// TIA Portal project "Tes simulation extract_V15.1" (V15.1) (continued)
VERSION : 0.1
   VAR_TEMP   // added for the SCL form of the ladder/FBD networks
      _w1 : Bool;
      _w2 : Bool;
   END_VAR
BEGIN

REGION Network 1: BUKA VALVE VP 1 DAN VP 5
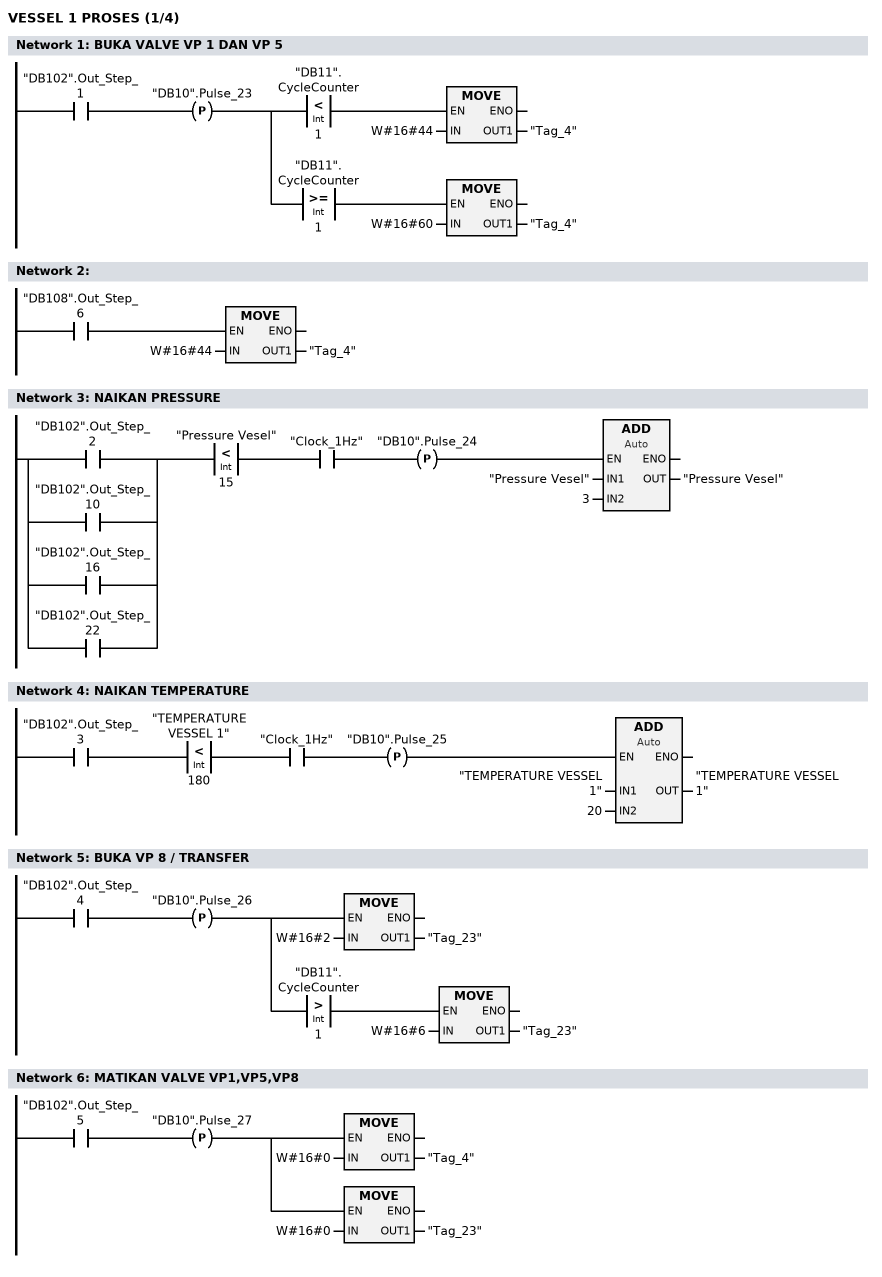
   RUNG wire#powerrail
      Contact( "DB102".Out_Step_1 )
      P_Trig( "DB10".Pulse_23 )
      wire#w1
      { S7_Templates := "SrcType := Int" } LT_Contact(in1 := "DB11".CycleCounter, in2 := 1)
      Move(in := W#16#44, out1 => "Tag_4")
   END_RUNG
   RUNG wire#w1
      { S7_Templates := "SrcType := Int" } GE_Contact(in1 := "DB11".CycleCounter, in2 := 1)
      Move(in := W#16#60, out1 => "Tag_4")
   END_RUNG
   // the same network as SCL:
   #_w1 := "DB102".Out_Step_1 AND NOT "DB10".Pulse_23;   // rising edge
   "DB10".Pulse_23 := "DB102".Out_Step_1;
   IF #_w1 AND ("DB11".CycleCounter < 1) THEN "Tag_4" := W#16#44; END_IF;
   IF #_w1 AND ("DB11".CycleCounter >= 1) THEN "Tag_4" := W#16#60; END_IF;
END_REGION

REGION Network 2
   RUNG wire#powerrail
      Contact( "DB108".Out_Step_6 )
      Move(in := W#16#44, out1 => "Tag_4")
   END_RUNG
   // the same network as SCL:
   IF "DB108".Out_Step_6 THEN "Tag_4" := W#16#44; END_IF;
END_REGION

REGION Network 3: NAIKAN PRESSURE
   RUNG wire#powerrail
      Contact( "DB102".Out_Step_2 )
      wire#w1
      { S7_Templates := "SrcType := Int" } LT_Contact(in1 := "Pressure Vesel", in2 := 15)
      Contact( "Clock_1Hz" )
      P_Trig( "DB10".Pulse_24 )
      Add(in1 := "Pressure Vesel", in2 := 3, out => "Pressure Vesel")
   END_RUNG
   RUNG wire#powerrail
      Contact( "DB102".Out_Step_10 )
   END_RUNG wire#w1
   RUNG wire#powerrail
      Contact( "DB102".Out_Step_16 )
   END_RUNG wire#w1
   RUNG wire#powerrail
      Contact( "DB102".Out_Step_22 )
   END_RUNG wire#w1
   // the same network as SCL:
   #_w1 := ("DB102".Out_Step_2 OR "DB102".Out_Step_10 OR "DB102".Out_Step_16 OR "DB102".Out_Step_22) AND ("Pressure Vesel" < 15) AND "Clock_1Hz";
   #_w2 := #_w1 AND NOT "DB10".Pulse_24;   // rising edge
   "DB10".Pulse_24 := #_w1;
   IF #_w2 THEN "Pressure Vesel" := "Pressure Vesel" + 3; END_IF;
END_REGION

REGION Network 4: NAIKAN TEMPERATURE
   RUNG wire#powerrail
      Contact( "DB102".Out_Step_3 )
      { S7_Templates := "SrcType := Int" } LT_Contact(in1 := "TEMPERATURE VESSEL 1", in2 := 180)
      Contact( "Clock_1Hz" )
      P_Trig( "DB10".Pulse_25 )
      Add(in1 := "TEMPERATURE VESSEL 1", in2 := 20, out => "TEMPERATURE VESSEL 1")
   END_RUNG
   // the same network as SCL:
   #_w1 := "DB102".Out_Step_3 AND ("TEMPERATURE VESSEL 1" < 180) AND "Clock_1Hz";
   #_w2 := #_w1 AND NOT "DB10".Pulse_25;   // rising edge
   "DB10".Pulse_25 := #_w1;
   IF #_w2 THEN "TEMPERATURE VESSEL 1" := "TEMPERATURE VESSEL 1" + 20; END_IF;
END_REGION

REGION Network 5: BUKA VP 8 / TRANSFER
   RUNG wire#powerrail
      Contact( "DB102".Out_Step_4 )
      P_Trig( "DB10".Pulse_26 )
      wire#w1
      Move(in := W#16#2, out1 => "Tag_23")
   END_RUNG
   RUNG wire#w1
      { S7_Templates := "SrcType := Int" } GT_Contact(in1 := "DB11".CycleCounter, in2 := 1)
      Move(in := W#16#6, out1 => "Tag_23")
   END_RUNG
   // the same network as SCL:
   #_w1 := "DB102".Out_Step_4 AND NOT "DB10".Pulse_26;   // rising edge
   "DB10".Pulse_26 := "DB102".Out_Step_4;
   IF #_w1 THEN "Tag_23" := W#16#2; END_IF;
   IF #_w1 AND ("DB11".CycleCounter > 1) THEN "Tag_23" := W#16#6; END_IF;
END_REGION

REGION Network 6: MATIKAN VALVE VP1,VP5,VP8
   RUNG wire#powerrail
      Contact( "DB102".Out_Step_5 )
      P_Trig( "DB10".Pulse_27 )
      wire#w1
      Move(in := W#16#0, out1 => "Tag_4")
   END_RUNG
   RUNG wire#w1
      Move(in := W#16#0, out1 => "Tag_23")
   END_RUNG
   // the same network as SCL:
   #_w1 := "DB102".Out_Step_5 AND NOT "DB10".Pulse_27;   // rising edge
   "DB10".Pulse_27 := "DB102".Out_Step_5;
   IF #_w1 THEN
       "Tag_4" := W#16#0;
       "Tag_23" := W#16#0;
   END_IF;
END_REGION

REGION Network 7: NYALAKAN VB1
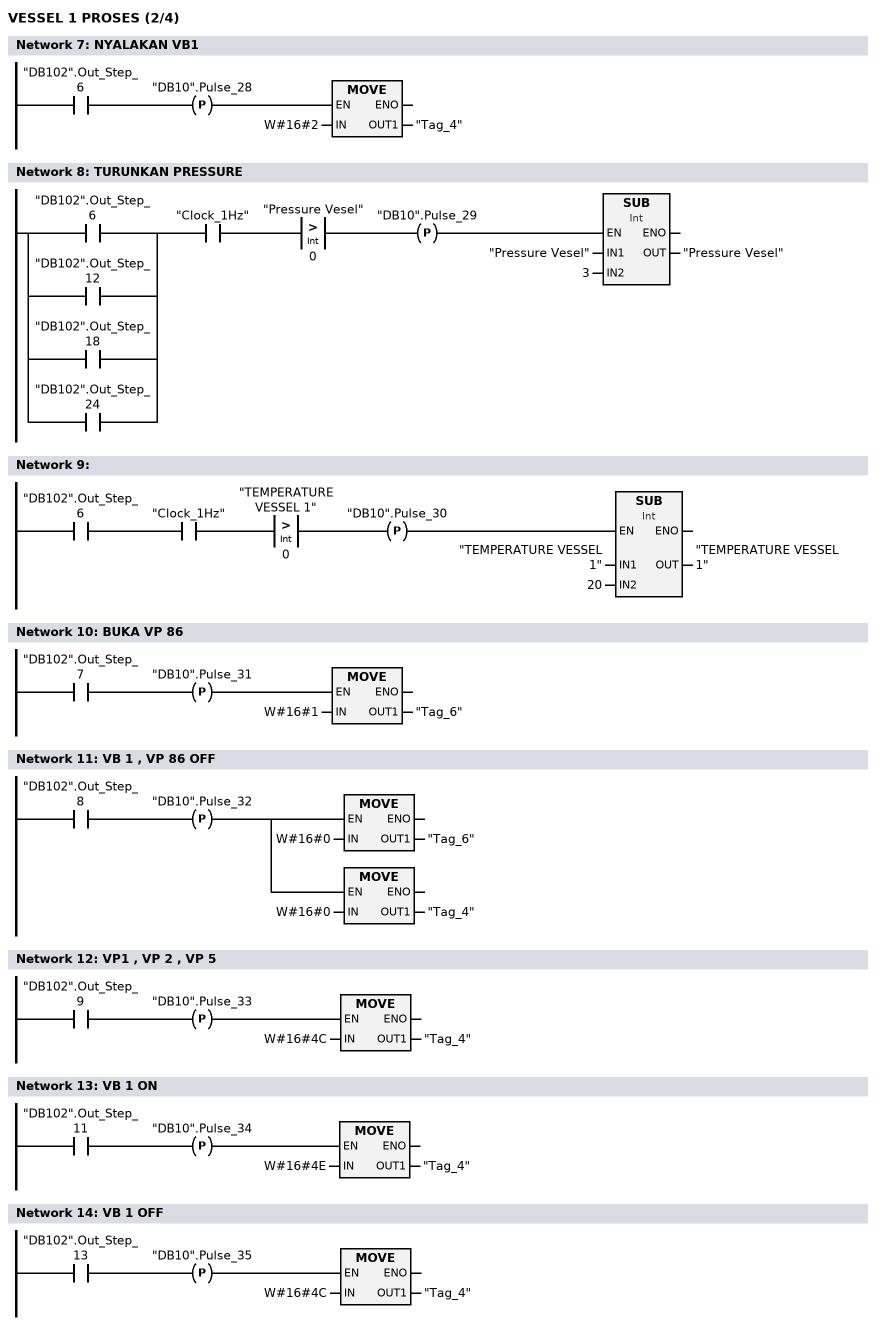
   RUNG wire#powerrail
      Contact( "DB102".Out_Step_6 )
      P_Trig( "DB10".Pulse_28 )
      Move(in := W#16#2, out1 => "Tag_4")
   END_RUNG
   // the same network as SCL:
   #_w1 := "DB102".Out_Step_6 AND NOT "DB10".Pulse_28;   // rising edge
   "DB10".Pulse_28 := "DB102".Out_Step_6;
   IF #_w1 THEN "Tag_4" := W#16#2; END_IF;
END_REGION

REGION Network 8: TURUNKAN PRESSURE
   RUNG wire#powerrail
      Contact( "DB102".Out_Step_6 )
      wire#w1
      Contact( "Clock_1Hz" )
      { S7_Templates := "SrcType := Int" } GT_Contact(in1 := "Pressure Vesel", in2 := 0)
      P_Trig( "DB10".Pulse_29 )
      { S7_Templates := "SrcType := Int" } Sub(in1 := "Pressure Vesel", in2 := 3, out => "Pressure Vesel")
   END_RUNG
   RUNG wire#powerrail
      Contact( "DB102".Out_Step_12 )
   END_RUNG wire#w1
   RUNG wire#powerrail
      Contact( "DB102".Out_Step_18 )
   END_RUNG wire#w1
   RUNG wire#powerrail
      Contact( "DB102".Out_Step_24 )
   END_RUNG wire#w1
   // the same network as SCL:
   #_w1 := ("DB102".Out_Step_6 OR "DB102".Out_Step_12 OR "DB102".Out_Step_18 OR "DB102".Out_Step_24) AND "Clock_1Hz" AND ("Pressure Vesel" > 0);
   #_w2 := #_w1 AND NOT "DB10".Pulse_29;   // rising edge
   "DB10".Pulse_29 := #_w1;
   IF #_w2 THEN "Pressure Vesel" := "Pressure Vesel" - 3; END_IF;
END_REGION

REGION Network 9
   RUNG wire#powerrail
      Contact( "DB102".Out_Step_6 )
      Contact( "Clock_1Hz" )
      { S7_Templates := "SrcType := Int" } GT_Contact(in1 := "TEMPERATURE VESSEL 1", in2 := 0)
      P_Trig( "DB10".Pulse_30 )
      { S7_Templates := "SrcType := Int" } Sub(in1 := "TEMPERATURE VESSEL 1", in2 := 20, out => "TEMPERATURE VESSEL 1")
   END_RUNG
   // the same network as SCL:
   #_w1 := "DB102".Out_Step_6 AND "Clock_1Hz" AND ("TEMPERATURE VESSEL 1" > 0);
   #_w2 := #_w1 AND NOT "DB10".Pulse_30;   // rising edge
   "DB10".Pulse_30 := #_w1;
   IF #_w2 THEN "TEMPERATURE VESSEL 1" := "TEMPERATURE VESSEL 1" - 20; END_IF;
END_REGION

REGION Network 10: BUKA VP 86
   RUNG wire#powerrail
      Contact( "DB102".Out_Step_7 )
      P_Trig( "DB10".Pulse_31 )
      Move(in := W#16#1, out1 => "Tag_6")
   END_RUNG
   // the same network as SCL:
   #_w1 := "DB102".Out_Step_7 AND NOT "DB10".Pulse_31;   // rising edge
   "DB10".Pulse_31 := "DB102".Out_Step_7;
   IF #_w1 THEN "Tag_6" := W#16#1; END_IF;
END_REGION

REGION Network 11: VB 1 , VP 86 OFF
   RUNG wire#powerrail
      Contact( "DB102".Out_Step_8 )
      P_Trig( "DB10".Pulse_32 )
      wire#w1
      Move(in := W#16#0, out1 => "Tag_6")
   END_RUNG
   RUNG wire#w1
      Move(in := W#16#0, out1 => "Tag_4")
   END_RUNG
   // the same network as SCL:
   #_w1 := "DB102".Out_Step_8 AND NOT "DB10".Pulse_32;   // rising edge
   "DB10".Pulse_32 := "DB102".Out_Step_8;
   IF #_w1 THEN
       "Tag_6" := W#16#0;
       "Tag_4" := W#16#0;
   END_IF;
END_REGION

REGION Network 12: VP1 , VP 2 , VP 5
   RUNG wire#powerrail
      Contact( "DB102".Out_Step_9 )
      P_Trig( "DB10".Pulse_33 )
      Move(in := W#16#4C, out1 => "Tag_4")
   END_RUNG
   // the same network as SCL:
   #_w1 := "DB102".Out_Step_9 AND NOT "DB10".Pulse_33;   // rising edge
   "DB10".Pulse_33 := "DB102".Out_Step_9;
   IF #_w1 THEN "Tag_4" := W#16#4C; END_IF;
END_REGION

REGION Network 13: VB 1 ON
   RUNG wire#powerrail
      Contact( "DB102".Out_Step_11 )
      P_Trig( "DB10".Pulse_34 )
      Move(in := W#16#4E, out1 => "Tag_4")
   END_RUNG
   // the same network as SCL:
   #_w1 := "DB102".Out_Step_11 AND NOT "DB10".Pulse_34;   // rising edge
   "DB10".Pulse_34 := "DB102".Out_Step_11;
   IF #_w1 THEN "Tag_4" := W#16#4E; END_IF;
END_REGION

REGION Network 14: VB 1 OFF
   RUNG wire#powerrail
      Contact( "DB102".Out_Step_13 )
      P_Trig( "DB10".Pulse_35 )
      Move(in := W#16#4C, out1 => "Tag_4")
   END_RUNG
   // the same network as SCL:
   #_w1 := "DB102".Out_Step_13 AND NOT "DB10".Pulse_35;   // rising edge
   "DB10".Pulse_35 := "DB102".Out_Step_13;
   IF #_w1 THEN "Tag_4" := W#16#4C; END_IF;
END_REGION

REGION Network 15: , VP 86 ON
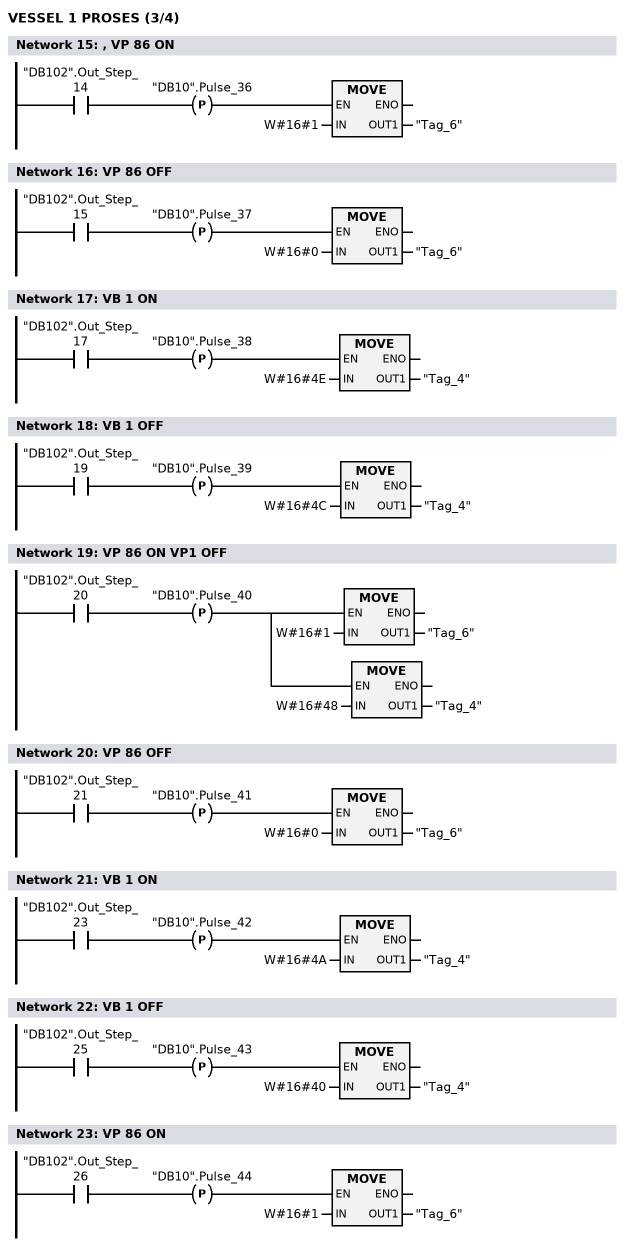
   RUNG wire#powerrail
      Contact( "DB102".Out_Step_14 )
      P_Trig( "DB10".Pulse_36 )
      Move(in := W#16#1, out1 => "Tag_6")
   END_RUNG
   // the same network as SCL:
   #_w1 := "DB102".Out_Step_14 AND NOT "DB10".Pulse_36;   // rising edge
   "DB10".Pulse_36 := "DB102".Out_Step_14;
   IF #_w1 THEN "Tag_6" := W#16#1; END_IF;
END_REGION

REGION Network 16: VP 86 OFF
   RUNG wire#powerrail
      Contact( "DB102".Out_Step_15 )
      P_Trig( "DB10".Pulse_37 )
      Move(in := W#16#0, out1 => "Tag_6")
   END_RUNG
   // the same network as SCL:
   #_w1 := "DB102".Out_Step_15 AND NOT "DB10".Pulse_37;   // rising edge
   "DB10".Pulse_37 := "DB102".Out_Step_15;
   IF #_w1 THEN "Tag_6" := W#16#0; END_IF;
END_REGION

REGION Network 17: VB 1 ON
   RUNG wire#powerrail
      Contact( "DB102".Out_Step_17 )
      P_Trig( "DB10".Pulse_38 )
      Move(in := W#16#4E, out1 => "Tag_4")
   END_RUNG
   // the same network as SCL:
   #_w1 := "DB102".Out_Step_17 AND NOT "DB10".Pulse_38;   // rising edge
   "DB10".Pulse_38 := "DB102".Out_Step_17;
   IF #_w1 THEN "Tag_4" := W#16#4E; END_IF;
END_REGION

REGION Network 18: VB 1 OFF
   RUNG wire#powerrail
      Contact( "DB102".Out_Step_19 )
      P_Trig( "DB10".Pulse_39 )
      Move(in := W#16#4C, out1 => "Tag_4")
   END_RUNG
   // the same network as SCL:
   #_w1 := "DB102".Out_Step_19 AND NOT "DB10".Pulse_39;   // rising edge
   "DB10".Pulse_39 := "DB102".Out_Step_19;
   IF #_w1 THEN "Tag_4" := W#16#4C; END_IF;
END_REGION

REGION Network 19: VP 86 ON VP1 OFF
   RUNG wire#powerrail
      Contact( "DB102".Out_Step_20 )
      P_Trig( "DB10".Pulse_40 )
      wire#w1
      Move(in := W#16#1, out1 => "Tag_6")
   END_RUNG
   RUNG wire#w1
      Move(in := W#16#48, out1 => "Tag_4")
   END_RUNG
   // the same network as SCL:
   #_w1 := "DB102".Out_Step_20 AND NOT "DB10".Pulse_40;   // rising edge
   "DB10".Pulse_40 := "DB102".Out_Step_20;
   IF #_w1 THEN
       "Tag_6" := W#16#1;
       "Tag_4" := W#16#48;
   END_IF;
END_REGION

REGION Network 20: VP 86 OFF
   RUNG wire#powerrail
      Contact( "DB102".Out_Step_21 )
      P_Trig( "DB10".Pulse_41 )
      Move(in := W#16#0, out1 => "Tag_6")
   END_RUNG
   // the same network as SCL:
   #_w1 := "DB102".Out_Step_21 AND NOT "DB10".Pulse_41;   // rising edge
   "DB10".Pulse_41 := "DB102".Out_Step_21;
   IF #_w1 THEN "Tag_6" := W#16#0; END_IF;
END_REGION

REGION Network 21: VB 1 ON
   RUNG wire#powerrail
      Contact( "DB102".Out_Step_23 )
      P_Trig( "DB10".Pulse_42 )
      Move(in := W#16#4A, out1 => "Tag_4")
   END_RUNG
   // the same network as SCL:
   #_w1 := "DB102".Out_Step_23 AND NOT "DB10".Pulse_42;   // rising edge
   "DB10".Pulse_42 := "DB102".Out_Step_23;
   IF #_w1 THEN "Tag_4" := W#16#4A; END_IF;
END_REGION

REGION Network 22: VB 1 OFF
   RUNG wire#powerrail
      Contact( "DB102".Out_Step_25 )
      P_Trig( "DB10".Pulse_43 )
      Move(in := W#16#40, out1 => "Tag_4")
   END_RUNG
   // the same network as SCL:
   #_w1 := "DB102".Out_Step_25 AND NOT "DB10".Pulse_43;   // rising edge
   "DB10".Pulse_43 := "DB102".Out_Step_25;
   IF #_w1 THEN "Tag_4" := W#16#40; END_IF;
END_REGION

REGION Network 23: VP 86 ON
   RUNG wire#powerrail
      Contact( "DB102".Out_Step_26 )
      P_Trig( "DB10".Pulse_44 )
      Move(in := W#16#1, out1 => "Tag_6")
   END_RUNG
   // the same network as SCL:
   #_w1 := "DB102".Out_Step_26 AND NOT "DB10".Pulse_44;   // rising edge
   "DB10".Pulse_44 := "DB102".Out_Step_26;
   IF #_w1 THEN "Tag_6" := W#16#1; END_IF;
END_REGION

REGION Network 24: VP 86 OFF VP 87 ON
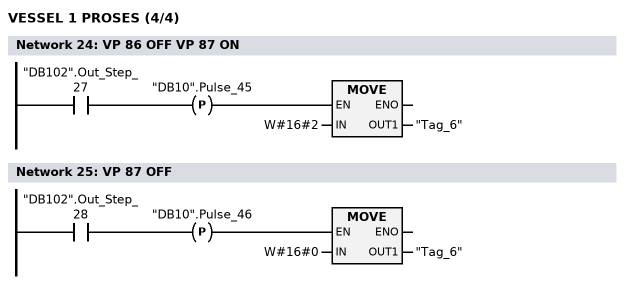
   RUNG wire#powerrail
      Contact( "DB102".Out_Step_27 )
      P_Trig( "DB10".Pulse_45 )
      Move(in := W#16#2, out1 => "Tag_6")
   END_RUNG
   // the same network as SCL:
   #_w1 := "DB102".Out_Step_27 AND NOT "DB10".Pulse_45;   // rising edge
   "DB10".Pulse_45 := "DB102".Out_Step_27;
   IF #_w1 THEN "Tag_6" := W#16#2; END_IF;
END_REGION

REGION Network 25: VP 87 OFF
   RUNG wire#powerrail
      Contact( "DB102".Out_Step_28 )
      P_Trig( "DB10".Pulse_46 )
      Move(in := W#16#0, out1 => "Tag_6")
   END_RUNG
   // the same network as SCL:
   #_w1 := "DB102".Out_Step_28 AND NOT "DB10".Pulse_46;   // rising edge
   "DB10".Pulse_46 := "DB102".Out_Step_28;
   IF #_w1 THEN "Tag_6" := W#16#0; END_IF;
END_REGION
END_FUNCTION

FUNCTION "SEQUENCE V1 PROSES" : Void   // FC7, LAD
{ S7_Optimized_Access := 'TRUE' }
VERSION : 0.1
   VAR_TEMP   // added for the SCL form of the ladder/FBD networks
      _w1 : Bool;
      _s5time1 : S5Time;
      _w2 : Bool;
      _w3 : Bool;
   END_VAR
BEGIN

REGION Network 1: START PROSES
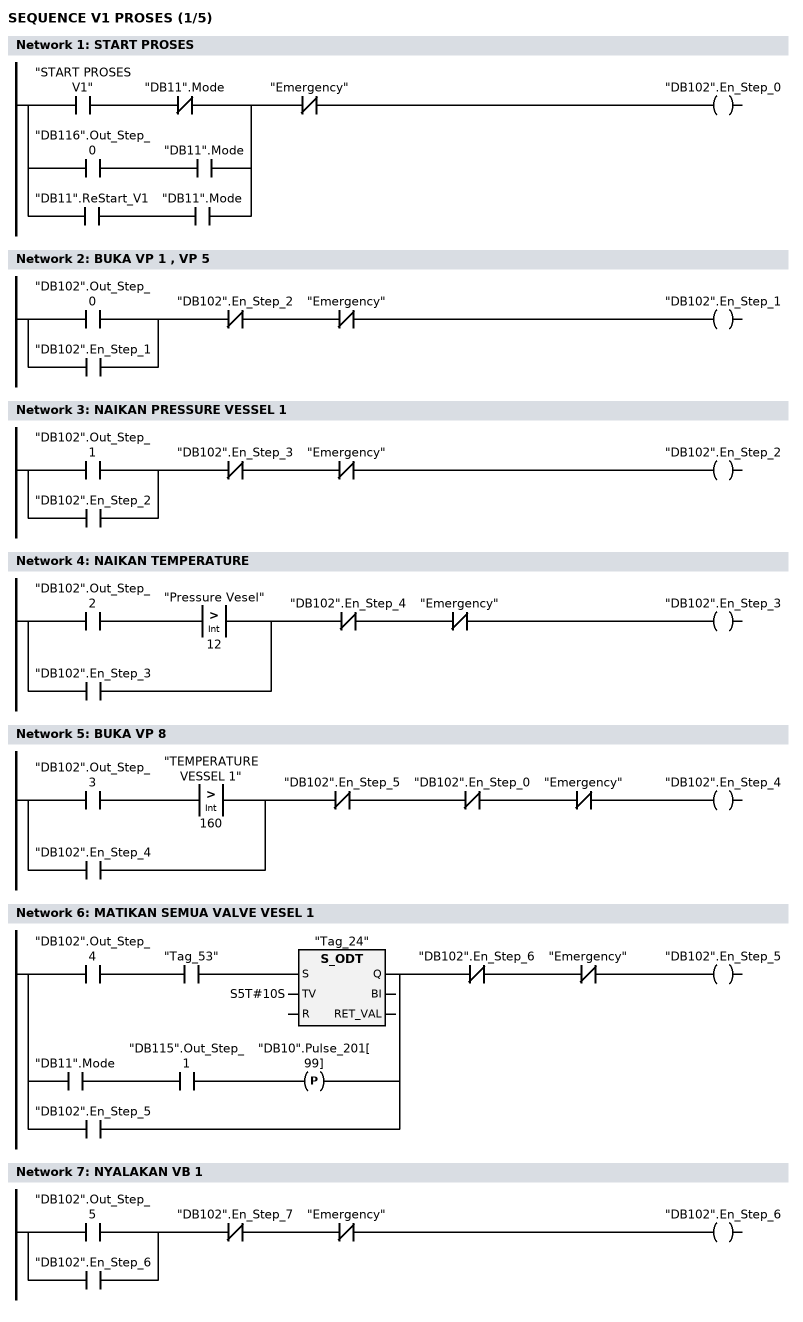
   RUNG wire#powerrail
      Contact( "START PROSES V1" )
      I_Contact( "DB11".Mode )
      wire#w1
      I_Contact( "Emergency" )
      Coil( "DB102".En_Step_0 )
   END_RUNG
   RUNG wire#powerrail
      Contact( "DB116".Out_Step_0 )
      Contact( "DB11".Mode )
   END_RUNG wire#w1
   RUNG wire#powerrail
      Contact( "DB11".ReStart_V1 )
      Contact( "DB11".Mode )
   END_RUNG wire#w1
   // the same network as SCL:
   "DB102".En_Step_0 := (("START PROSES V1" AND NOT "DB11".Mode) OR ("DB116".Out_Step_0 AND "DB11".Mode) OR ("DB11".ReStart_V1 AND "DB11".Mode)) AND NOT "Emergency";
END_REGION

REGION Network 2: BUKA VP 1 , VP 5
   RUNG wire#powerrail
      Contact( "DB102".Out_Step_0 )
      wire#w1
      I_Contact( "DB102".En_Step_2 )
      I_Contact( "Emergency" )
      Coil( "DB102".En_Step_1 )
   END_RUNG
   RUNG wire#powerrail
      Contact( "DB102".En_Step_1 )
   END_RUNG wire#w1
   // the same network as SCL:
   "DB102".En_Step_1 := ("DB102".Out_Step_0 OR "DB102".En_Step_1) AND NOT "DB102".En_Step_2 AND NOT "Emergency";
END_REGION

REGION Network 3: NAIKAN PRESSURE VESSEL 1
   RUNG wire#powerrail
      Contact( "DB102".Out_Step_1 )
      wire#w1
      I_Contact( "DB102".En_Step_3 )
      I_Contact( "Emergency" )
      Coil( "DB102".En_Step_2 )
   END_RUNG
   RUNG wire#powerrail
      Contact( "DB102".En_Step_2 )
   END_RUNG wire#w1
   // the same network as SCL:
   "DB102".En_Step_2 := ("DB102".Out_Step_1 OR "DB102".En_Step_2) AND NOT "DB102".En_Step_3 AND NOT "Emergency";
END_REGION

REGION Network 4: NAIKAN TEMPERATURE
   RUNG wire#powerrail
      Contact( "DB102".Out_Step_2 )
      { S7_Templates := "SrcType := Int" } GT_Contact(in1 := "Pressure Vesel", in2 := 12)
      wire#w1
      I_Contact( "DB102".En_Step_4 )
      I_Contact( "Emergency" )
      Coil( "DB102".En_Step_3 )
   END_RUNG
   RUNG wire#powerrail
      Contact( "DB102".En_Step_3 )
   END_RUNG wire#w1
   // the same network as SCL:
   "DB102".En_Step_3 := (("DB102".Out_Step_2 AND ("Pressure Vesel" > 12)) OR "DB102".En_Step_3) AND NOT "DB102".En_Step_4 AND NOT "Emergency";
END_REGION

REGION Network 5: BUKA VP 8
   RUNG wire#powerrail
      Contact( "DB102".Out_Step_3 )
      { S7_Templates := "SrcType := Int" } GT_Contact(in1 := "TEMPERATURE VESSEL 1", in2 := 160)
      wire#w1
      I_Contact( "DB102".En_Step_5 )
      I_Contact( "DB102".En_Step_0 )
      I_Contact( "Emergency" )
      Coil( "DB102".En_Step_4 )
   END_RUNG
   RUNG wire#powerrail
      Contact( "DB102".En_Step_4 )
   END_RUNG wire#w1
   // the same network as SCL:
   "DB102".En_Step_4 := (("DB102".Out_Step_3 AND ("TEMPERATURE VESSEL 1" > 160)) OR "DB102".En_Step_4) AND NOT "DB102".En_Step_5 AND NOT "DB102".En_Step_0 AND NOT "Emergency";
END_REGION

REGION Network 6: MATIKAN SEMUA VALVE VESEL 1
   RUNG wire#powerrail
      Contact( "DB102".Out_Step_4 )
      Contact( "Tag_53" )
      S_ODT(T_NO := "Tag_24", TV := S5T#10S, R :=, BI =>, RET_VAL =>)
      wire#w1
      I_Contact( "DB102".En_Step_6 )
      I_Contact( "Emergency" )
      Coil( "DB102".En_Step_5 )
   END_RUNG
   RUNG wire#powerrail
      Contact( "DB11".Mode )
      Contact( "DB115".Out_Step_1 )
      P_Trig( "DB10".Pulse_201[99] )
   END_RUNG wire#w1
   RUNG wire#powerrail
      Contact( "DB102".En_Step_5 )
   END_RUNG wire#w1
   // the same network as SCL:
   #_s5time1 := S_ODT(T_NO := "Tag_24", S := "DB102".Out_Step_4 AND "Tag_53", TV := S5T#10S, Q => #_w1);
   #_w2 := "DB11".Mode AND "DB115".Out_Step_1;
   #_w3 := #_w2 AND NOT "DB10".Pulse_201[99];   // rising edge
   "DB10".Pulse_201[99] := #_w2;
   "DB102".En_Step_5 := (#_w1 OR #_w3 OR "DB102".En_Step_5) AND NOT "DB102".En_Step_6 AND NOT "Emergency";
END_REGION

REGION Network 7: NYALAKAN VB 1
   RUNG wire#powerrail
      Contact( "DB102".Out_Step_5 )
      wire#w1
      I_Contact( "DB102".En_Step_7 )
      I_Contact( "Emergency" )
      Coil( "DB102".En_Step_6 )
   END_RUNG
   RUNG wire#powerrail
      Contact( "DB102".En_Step_6 )
   END_RUNG wire#w1
   // the same network as SCL:
   "DB102".En_Step_6 := ("DB102".Out_Step_5 OR "DB102".En_Step_6) AND NOT "DB102".En_Step_7 AND NOT "Emergency";
END_REGION

REGION Network 8
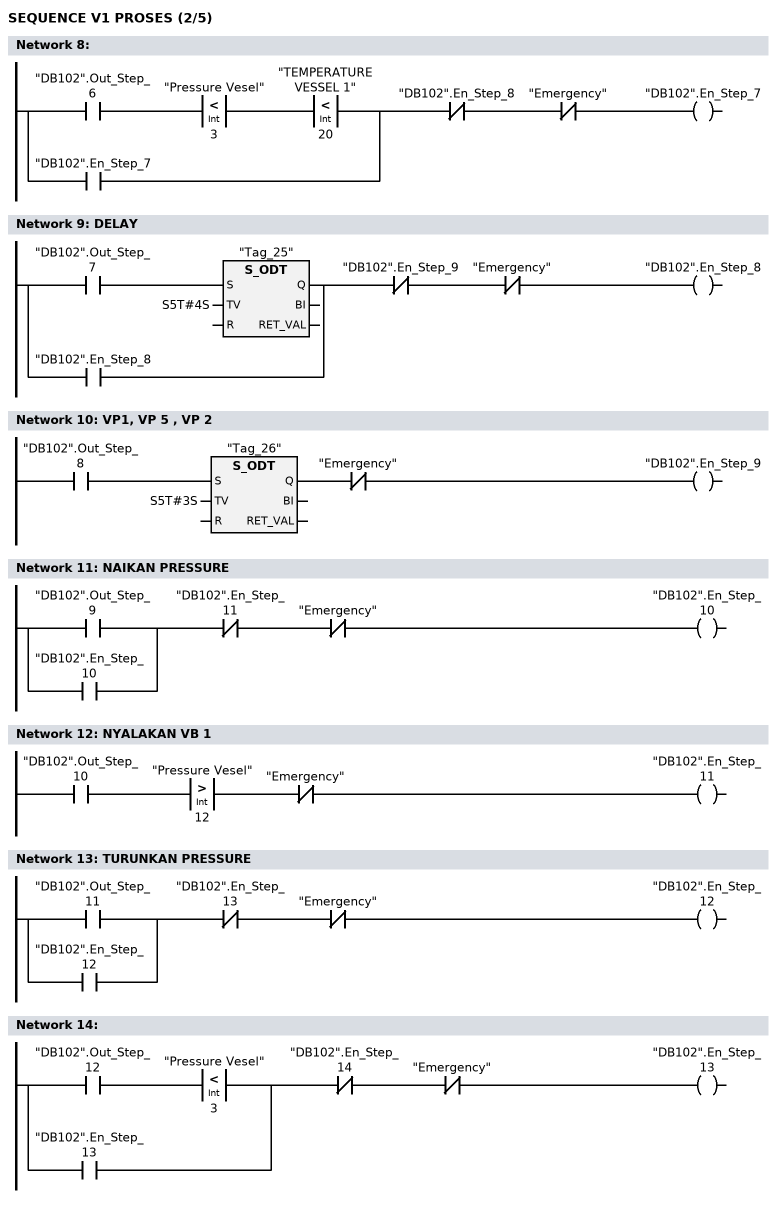
   RUNG wire#powerrail
      Contact( "DB102".Out_Step_6 )
      { S7_Templates := "SrcType := Int" } LT_Contact(in1 := "Pressure Vesel", in2 := 3)
      { S7_Templates := "SrcType := Int" } LT_Contact(in1 := "TEMPERATURE VESSEL 1", in2 := 20)
      wire#w1
      I_Contact( "DB102".En_Step_8 )
      I_Contact( "Emergency" )
      Coil( "DB102".En_Step_7 )
   END_RUNG
   RUNG wire#powerrail
      Contact( "DB102".En_Step_7 )
   END_RUNG wire#w1
   // the same network as SCL:
   "DB102".En_Step_7 := (("DB102".Out_Step_6 AND ("Pressure Vesel" < 3) AND ("TEMPERATURE VESSEL 1" < 20)) OR "DB102".En_Step_7) AND NOT "DB102".En_Step_8 AND NOT "Emergency";
END_REGION

REGION Network 9: DELAY
   RUNG wire#powerrail
      Contact( "DB102".Out_Step_7 )
      S_ODT(T_NO := "Tag_25", TV := S5T#4S, R :=, BI =>, RET_VAL =>)
      wire#w1
      I_Contact( "DB102".En_Step_9 )
      I_Contact( "Emergency" )
      Coil( "DB102".En_Step_8 )
   END_RUNG
   RUNG wire#powerrail
      Contact( "DB102".En_Step_8 )
   END_RUNG wire#w1
   // the same network as SCL:
   #_s5time1 := S_ODT(T_NO := "Tag_25", S := "DB102".Out_Step_7, TV := S5T#4S, Q => #_w1);
   "DB102".En_Step_8 := (#_w1 OR "DB102".En_Step_8) AND NOT "DB102".En_Step_9 AND NOT "Emergency";
END_REGION

REGION Network 10: VP1, VP 5 , VP 2
   RUNG wire#powerrail
      Contact( "DB102".Out_Step_8 )
      S_ODT(T_NO := "Tag_26", TV := S5T#3S, R :=, BI =>, RET_VAL =>)
      I_Contact( "Emergency" )
      Coil( "DB102".En_Step_9 )
   END_RUNG
   // the same network as SCL:
   #_s5time1 := S_ODT(T_NO := "Tag_26", S := "DB102".Out_Step_8, TV := S5T#3S, Q => #_w1);
   "DB102".En_Step_9 := #_w1 AND NOT "Emergency";
END_REGION

REGION Network 11: NAIKAN PRESSURE
   RUNG wire#powerrail
      Contact( "DB102".Out_Step_9 )
      wire#w1
      I_Contact( "DB102".En_Step_11 )
      I_Contact( "Emergency" )
      Coil( "DB102".En_Step_10 )
   END_RUNG
   RUNG wire#powerrail
      Contact( "DB102".En_Step_10 )
   END_RUNG wire#w1
   // the same network as SCL:
   "DB102".En_Step_10 := ("DB102".Out_Step_9 OR "DB102".En_Step_10) AND NOT "DB102".En_Step_11 AND NOT "Emergency";
END_REGION

REGION Network 12: NYALAKAN VB 1
   RUNG wire#powerrail
      Contact( "DB102".Out_Step_10 )
      { S7_Templates := "SrcType := Int" } GT_Contact(in1 := "Pressure Vesel", in2 := 12)
      I_Contact( "Emergency" )
      Coil( "DB102".En_Step_11 )
   END_RUNG
   // the same network as SCL:
   "DB102".En_Step_11 := "DB102".Out_Step_10 AND ("Pressure Vesel" > 12) AND NOT "Emergency";
END_REGION

REGION Network 13: TURUNKAN PRESSURE
   RUNG wire#powerrail
      Contact( "DB102".Out_Step_11 )
      wire#w1
      I_Contact( "DB102".En_Step_13 )
      I_Contact( "Emergency" )
      Coil( "DB102".En_Step_12 )
   END_RUNG
   RUNG wire#powerrail
      Contact( "DB102".En_Step_12 )
   END_RUNG wire#w1
   // the same network as SCL:
   "DB102".En_Step_12 := ("DB102".Out_Step_11 OR "DB102".En_Step_12) AND NOT "DB102".En_Step_13 AND NOT "Emergency";
END_REGION

REGION Network 14
   RUNG wire#powerrail
      Contact( "DB102".Out_Step_12 )
      { S7_Templates := "SrcType := Int" } LT_Contact(in1 := "Pressure Vesel", in2 := 3)
      wire#w1
      I_Contact( "DB102".En_Step_14 )
      I_Contact( "Emergency" )
      Coil( "DB102".En_Step_13 )
   END_RUNG
   RUNG wire#powerrail
      Contact( "DB102".En_Step_13 )
   END_RUNG wire#w1
   // the same network as SCL:
   "DB102".En_Step_13 := (("DB102".Out_Step_12 AND ("Pressure Vesel" < 3)) OR "DB102".En_Step_13) AND NOT "DB102".En_Step_14 AND NOT "Emergency";
END_REGION

REGION Network 15
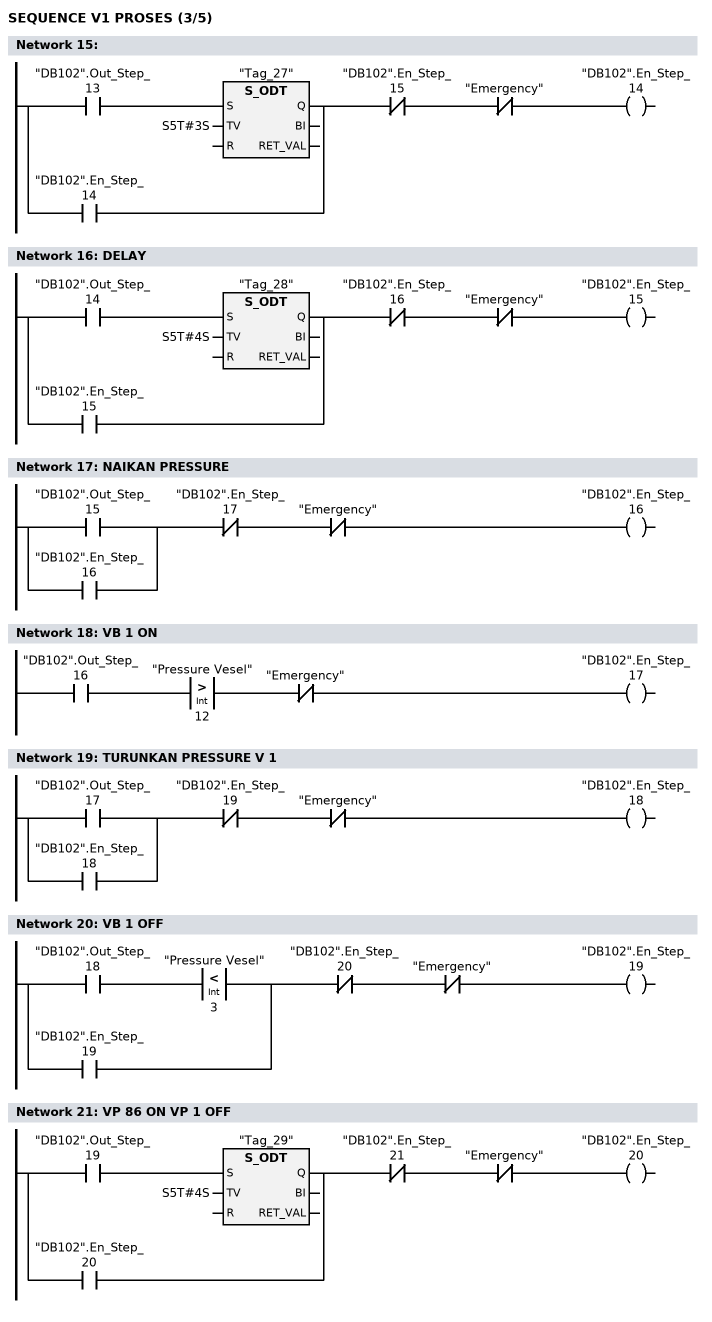
   RUNG wire#powerrail
      Contact( "DB102".Out_Step_13 )
      S_ODT(T_NO := "Tag_27", TV := S5T#3S, R :=, BI =>, RET_VAL =>)
      wire#w1
      I_Contact( "DB102".En_Step_15 )
      I_Contact( "Emergency" )
      Coil( "DB102".En_Step_14 )
   END_RUNG
   RUNG wire#powerrail
      Contact( "DB102".En_Step_14 )
   END_RUNG wire#w1
   // the same network as SCL:
   #_s5time1 := S_ODT(T_NO := "Tag_27", S := "DB102".Out_Step_13, TV := S5T#3S, Q => #_w1);
   "DB102".En_Step_14 := (#_w1 OR "DB102".En_Step_14) AND NOT "DB102".En_Step_15 AND NOT "Emergency";
END_REGION

REGION Network 16: DELAY
   RUNG wire#powerrail
      Contact( "DB102".Out_Step_14 )
      S_ODT(T_NO := "Tag_28", TV := S5T#4S, R :=, BI =>, RET_VAL =>)
      wire#w1
      I_Contact( "DB102".En_Step_16 )
      I_Contact( "Emergency" )
      Coil( "DB102".En_Step_15 )
   END_RUNG
   RUNG wire#powerrail
      Contact( "DB102".En_Step_15 )
   END_RUNG wire#w1
   // the same network as SCL:
   #_s5time1 := S_ODT(T_NO := "Tag_28", S := "DB102".Out_Step_14, TV := S5T#4S, Q => #_w1);
   "DB102".En_Step_15 := (#_w1 OR "DB102".En_Step_15) AND NOT "DB102".En_Step_16 AND NOT "Emergency";
END_REGION

REGION Network 17: NAIKAN PRESSURE
   RUNG wire#powerrail
      Contact( "DB102".Out_Step_15 )
      wire#w1
      I_Contact( "DB102".En_Step_17 )
      I_Contact( "Emergency" )
      Coil( "DB102".En_Step_16 )
   END_RUNG
   RUNG wire#powerrail
      Contact( "DB102".En_Step_16 )
   END_RUNG wire#w1
   // the same network as SCL:
   "DB102".En_Step_16 := ("DB102".Out_Step_15 OR "DB102".En_Step_16) AND NOT "DB102".En_Step_17 AND NOT "Emergency";
END_REGION

REGION Network 18: VB 1 ON
   RUNG wire#powerrail
      Contact( "DB102".Out_Step_16 )
      { S7_Templates := "SrcType := Int" } GT_Contact(in1 := "Pressure Vesel", in2 := 12)
      I_Contact( "Emergency" )
      Coil( "DB102".En_Step_17 )
   END_RUNG
   // the same network as SCL:
   "DB102".En_Step_17 := "DB102".Out_Step_16 AND ("Pressure Vesel" > 12) AND NOT "Emergency";
END_REGION

REGION Network 19: TURUNKAN PRESSURE V 1
   RUNG wire#powerrail
      Contact( "DB102".Out_Step_17 )
      wire#w1
      I_Contact( "DB102".En_Step_19 )
      I_Contact( "Emergency" )
      Coil( "DB102".En_Step_18 )
   END_RUNG
   RUNG wire#powerrail
      Contact( "DB102".En_Step_18 )
   END_RUNG wire#w1
   // the same network as SCL:
   "DB102".En_Step_18 := ("DB102".Out_Step_17 OR "DB102".En_Step_18) AND NOT "DB102".En_Step_19 AND NOT "Emergency";
END_REGION

REGION Network 20: VB 1 OFF
   RUNG wire#powerrail
      Contact( "DB102".Out_Step_18 )
      { S7_Templates := "SrcType := Int" } LT_Contact(in1 := "Pressure Vesel", in2 := 3)
      wire#w1
      I_Contact( "DB102".En_Step_20 )
      I_Contact( "Emergency" )
      Coil( "DB102".En_Step_19 )
   END_RUNG
   RUNG wire#powerrail
      Contact( "DB102".En_Step_19 )
   END_RUNG wire#w1
   // the same network as SCL:
   "DB102".En_Step_19 := (("DB102".Out_Step_18 AND ("Pressure Vesel" < 3)) OR "DB102".En_Step_19) AND NOT "DB102".En_Step_20 AND NOT "Emergency";
END_REGION

REGION Network 21: VP 86 ON VP 1 OFF
   RUNG wire#powerrail
      Contact( "DB102".Out_Step_19 )
      S_ODT(T_NO := "Tag_29", TV := S5T#4S, R :=, BI =>, RET_VAL =>)
      wire#w1
      I_Contact( "DB102".En_Step_21 )
      I_Contact( "Emergency" )
      Coil( "DB102".En_Step_20 )
   END_RUNG
   RUNG wire#powerrail
      Contact( "DB102".En_Step_20 )
   END_RUNG wire#w1
   // the same network as SCL:
   #_s5time1 := S_ODT(T_NO := "Tag_29", S := "DB102".Out_Step_19, TV := S5T#4S, Q => #_w1);
   "DB102".En_Step_20 := (#_w1 OR "DB102".En_Step_20) AND NOT "DB102".En_Step_21 AND NOT "Emergency";
END_REGION

REGION Network 22: VP 86 OFF VP 87 ON
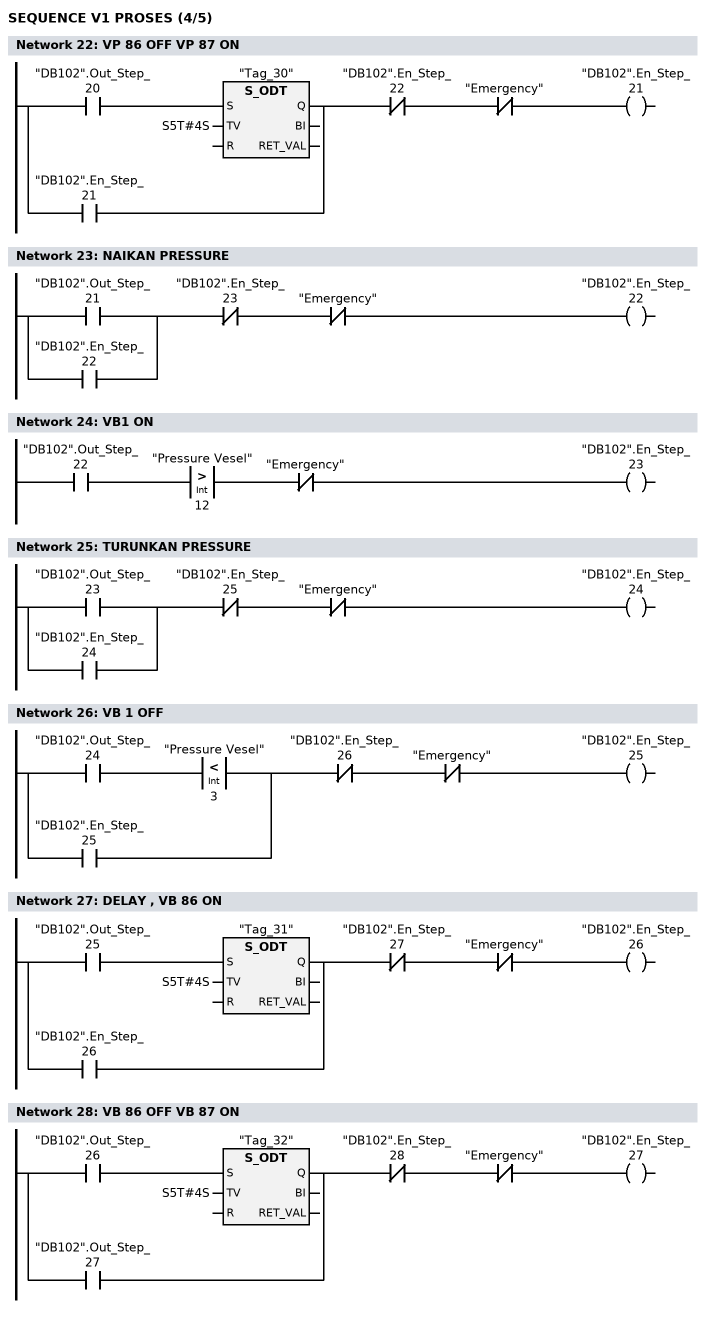
   RUNG wire#powerrail
      Contact( "DB102".Out_Step_20 )
      S_ODT(T_NO := "Tag_30", TV := S5T#4S, R :=, BI =>, RET_VAL =>)
      wire#w1
      I_Contact( "DB102".En_Step_22 )
      I_Contact( "Emergency" )
      Coil( "DB102".En_Step_21 )
   END_RUNG
   RUNG wire#powerrail
      Contact( "DB102".En_Step_21 )
   END_RUNG wire#w1
   // the same network as SCL:
   #_s5time1 := S_ODT(T_NO := "Tag_30", S := "DB102".Out_Step_20, TV := S5T#4S, Q => #_w1);
   "DB102".En_Step_21 := (#_w1 OR "DB102".En_Step_21) AND NOT "DB102".En_Step_22 AND NOT "Emergency";
END_REGION

REGION Network 23: NAIKAN PRESSURE
   RUNG wire#powerrail
      Contact( "DB102".Out_Step_21 )
      wire#w1
      I_Contact( "DB102".En_Step_23 )
      I_Contact( "Emergency" )
      Coil( "DB102".En_Step_22 )
   END_RUNG
   RUNG wire#powerrail
      Contact( "DB102".En_Step_22 )
   END_RUNG wire#w1
   // the same network as SCL:
   "DB102".En_Step_22 := ("DB102".Out_Step_21 OR "DB102".En_Step_22) AND NOT "DB102".En_Step_23 AND NOT "Emergency";
END_REGION

REGION Network 24: VB1 ON
   RUNG wire#powerrail
      Contact( "DB102".Out_Step_22 )
      { S7_Templates := "SrcType := Int" } GT_Contact(in1 := "Pressure Vesel", in2 := 12)
      I_Contact( "Emergency" )
      Coil( "DB102".En_Step_23 )
   END_RUNG
   // the same network as SCL:
   "DB102".En_Step_23 := "DB102".Out_Step_22 AND ("Pressure Vesel" > 12) AND NOT "Emergency";
END_REGION

REGION Network 25: TURUNKAN PRESSURE
   RUNG wire#powerrail
      Contact( "DB102".Out_Step_23 )
      wire#w1
      I_Contact( "DB102".En_Step_25 )
      I_Contact( "Emergency" )
      Coil( "DB102".En_Step_24 )
   END_RUNG
   RUNG wire#powerrail
      Contact( "DB102".En_Step_24 )
   END_RUNG wire#w1
   // the same network as SCL:
   "DB102".En_Step_24 := ("DB102".Out_Step_23 OR "DB102".En_Step_24) AND NOT "DB102".En_Step_25 AND NOT "Emergency";
END_REGION

REGION Network 26: VB 1 OFF
   RUNG wire#powerrail
      Contact( "DB102".Out_Step_24 )
      { S7_Templates := "SrcType := Int" } LT_Contact(in1 := "Pressure Vesel", in2 := 3)
      wire#w1
      I_Contact( "DB102".En_Step_26 )
      I_Contact( "Emergency" )
      Coil( "DB102".En_Step_25 )
   END_RUNG
   RUNG wire#powerrail
      Contact( "DB102".En_Step_25 )
   END_RUNG wire#w1
   // the same network as SCL:
   "DB102".En_Step_25 := (("DB102".Out_Step_24 AND ("Pressure Vesel" < 3)) OR "DB102".En_Step_25) AND NOT "DB102".En_Step_26 AND NOT "Emergency";
END_REGION

REGION Network 27: DELAY , VB 86 ON
   RUNG wire#powerrail
      Contact( "DB102".Out_Step_25 )
      S_ODT(T_NO := "Tag_31", TV := S5T#4S, R :=, BI =>, RET_VAL =>)
      wire#w1
      I_Contact( "DB102".En_Step_27 )
      I_Contact( "Emergency" )
      Coil( "DB102".En_Step_26 )
   END_RUNG
   RUNG wire#powerrail
      Contact( "DB102".En_Step_26 )
   END_RUNG wire#w1
   // the same network as SCL:
   #_s5time1 := S_ODT(T_NO := "Tag_31", S := "DB102".Out_Step_25, TV := S5T#4S, Q => #_w1);
   "DB102".En_Step_26 := (#_w1 OR "DB102".En_Step_26) AND NOT "DB102".En_Step_27 AND NOT "Emergency";
END_REGION

REGION Network 28: VB 86 OFF VB 87 ON
   RUNG wire#powerrail
      Contact( "DB102".Out_Step_26 )
      S_ODT(T_NO := "Tag_32", TV := S5T#4S, R :=, BI =>, RET_VAL =>)
      wire#w1
      I_Contact( "DB102".En_Step_28 )
      I_Contact( "Emergency" )
      Coil( "DB102".En_Step_27 )
   END_RUNG
   RUNG wire#powerrail
      Contact( "DB102".Out_Step_27 )
   END_RUNG wire#w1
   // the same network as SCL:
   #_s5time1 := S_ODT(T_NO := "Tag_32", S := "DB102".Out_Step_26, TV := S5T#4S, Q => #_w1);
   "DB102".En_Step_27 := (#_w1 OR "DB102".Out_Step_27) AND NOT "DB102".En_Step_28 AND NOT "Emergency";
END_REGION

REGION Network 29
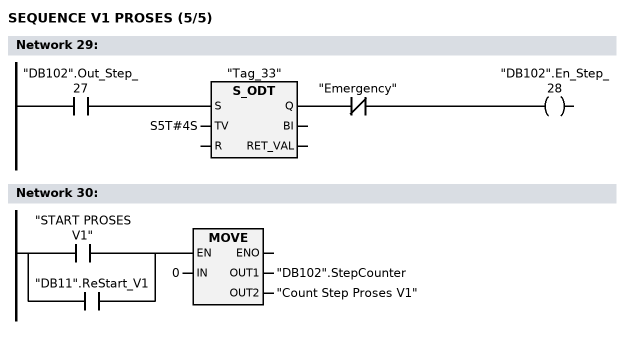
   RUNG wire#powerrail
      Contact( "DB102".Out_Step_27 )
      S_ODT(T_NO := "Tag_33", TV := S5T#4S, R :=, BI =>, RET_VAL =>)
      I_Contact( "Emergency" )
      Coil( "DB102".En_Step_28 )
   END_RUNG
   // the same network as SCL:
   #_s5time1 := S_ODT(T_NO := "Tag_33", S := "DB102".Out_Step_27, TV := S5T#4S, Q => #_w1);
   "DB102".En_Step_28 := #_w1 AND NOT "Emergency";
END_REGION

REGION Network 30
   RUNG wire#powerrail
      Contact( "START PROSES V1" )
      wire#w1
      Move(in := 0, out1 => "DB102".StepCounter, out2 => "Count Step Proses V1")
   END_RUNG
   RUNG wire#powerrail
      Contact( "DB11".ReStart_V1 )
   END_RUNG wire#w1
   // the same network as SCL:
   IF "START PROSES V1" OR "DB11".ReStart_V1 THEN
       "DB102".StepCounter := 0;
       "Count Step Proses V1" := 0;
   END_IF;
END_REGION
END_FUNCTION

FUNCTION "TRANSFER" : Void   // FC8, LAD
{ S7_Optimized_Access := 'TRUE' }
VERSION : 0.1
BEGIN

REGION Network 1
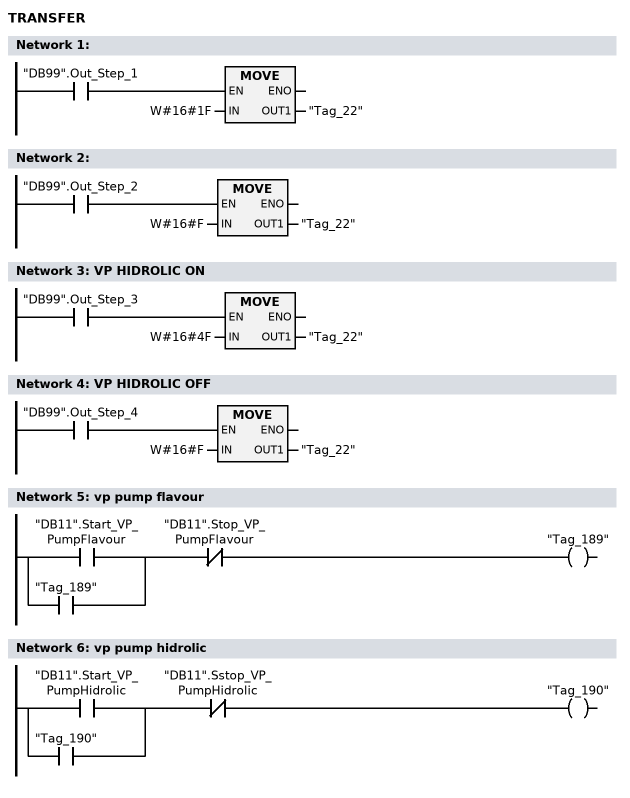
   RUNG wire#powerrail
      Contact( "DB99".Out_Step_1 )
      Move(in := W#16#1F, out1 => "Tag_22")
   END_RUNG
   // the same network as SCL:
   IF "DB99".Out_Step_1 THEN "Tag_22" := W#16#1F; END_IF;
END_REGION

REGION Network 2
   RUNG wire#powerrail
      Contact( "DB99".Out_Step_2 )
      Move(in := W#16#F, out1 => "Tag_22")
   END_RUNG
   // the same network as SCL:
   IF "DB99".Out_Step_2 THEN "Tag_22" := W#16#F; END_IF;
END_REGION

REGION Network 3: VP HIDROLIC ON
   RUNG wire#powerrail
      Contact( "DB99".Out_Step_3 )
      Move(in := W#16#4F, out1 => "Tag_22")
   END_RUNG
   // the same network as SCL:
   IF "DB99".Out_Step_3 THEN "Tag_22" := W#16#4F; END_IF;
END_REGION

REGION Network 4: VP HIDROLIC OFF
   RUNG wire#powerrail
      Contact( "DB99".Out_Step_4 )
      Move(in := W#16#F, out1 => "Tag_22")
   END_RUNG
   // the same network as SCL:
   IF "DB99".Out_Step_4 THEN "Tag_22" := W#16#F; END_IF;
END_REGION

REGION Network 5: vp pump flavour
   RUNG wire#powerrail
      Contact( "DB11".Start_VP_PumpFlavour )
      wire#w1
      I_Contact( "DB11".Stop_VP_PumpFlavour )
      Coil( "Tag_189" )
   END_RUNG
   RUNG wire#powerrail
      Contact( "Tag_189" )
   END_RUNG wire#w1
   // the same network as SCL:
   "Tag_189" := ("DB11".Start_VP_PumpFlavour OR "Tag_189") AND NOT "DB11".Stop_VP_PumpFlavour;
END_REGION

REGION Network 6: vp pump hidrolic
   RUNG wire#powerrail
      Contact( "DB11".Start_VP_PumpHidrolic )
      wire#w1
      I_Contact( "DB11".Sstop_VP_PumpHidrolic )
      Coil( "Tag_190" )
   END_RUNG
   RUNG wire#powerrail
      Contact( "Tag_190" )
   END_RUNG wire#w1
   // the same network as SCL:
   "Tag_190" := ("DB11".Start_VP_PumpHidrolic OR "Tag_190") AND NOT "DB11".Sstop_VP_PumpHidrolic;
END_REGION
END_FUNCTION

